// TIA Portal project "Project maybe not work 1.0" (V17) (continued)
REGION Network 7: Step 25 resetting the alarms
   "Data_Block_Reset_Seq".SeqStep[27] := "Data_Block_Reset_Seq".StepNumber = 27;
   "Data_Block_Reset_Seq".SeqConditions[27] := ("Data_Block_Reset_Seq".StepNumber = 27) AND NOT "FS-313.I" AND NOT "FS-214-I" AND "FS-213.I" AND NOT "FS-115.I" AND "FS-114.I" AND NOT "FS-113.I" AND NOT "FS-212.I" AND "HZ-413.I" AND NOT "Fire Alarm" AND NOT "QE-116.I" AND "QE-316.I";
   "Data_Block_Reset_Seq".SeqTimer[27].TON(IN := ("Data_Block_Reset_Seq".StepNumber = 27) AND (("FS-314.I" AND NOT "FS-315.I") OR (NOT "FS-315.I" AND NOT "FS-314.I")) AND NOT "FS-315.I" AND "Data_Block_Reset_Seq".SeqConditions[27],
                           PT := T#50MS);
   IF "Data_Block_Reset_Seq".SeqTimer[27].Q THEN
       "FCS-311.O" := FALSE;
       "FCS-312.O" := TRUE;
   END_IF;
   #_w1 := "Data_Block_Reset_Seq".StepNumber = 27;
   IF "Data_Block_Reset_Seq".SeqTimer[27].Q THEN "Data_Block_Reset_Seq".StepNumber := 28; END_IF;
   "Data_Block_Reset_Seq".SeqTimer_1[89].TON(IN := #_w1 AND NOT "FS-314.I" AND "FS-315.I" AND "Data_Block_Reset_Seq".SeqConditions[27],
                           PT := T#50MS);
   IF "Data_Block_Reset_Seq".SeqTimer_1[89].Q THEN "Data_Block_Reset_Seq".StepNumber := 28; END_IF;
END_REGION

REGION Network 8: Step 25 resetting the alarms
   "Data_Block_Reset_Seq".SeqStep[28] := "Data_Block_Reset_Seq".StepNumber = 28;
   "Data_Block_Reset_Seq".SeqConditions[28] := ("Data_Block_Reset_Seq".StepNumber = 28) AND NOT "FS-314.I" AND "FS-315.I" AND NOT "FS-313.I" AND NOT "FS-214-I" AND "FS-213.I" AND NOT "FS-115.I" AND "FS-114.I" AND NOT "FS-113.I" AND NOT "FS-212.I" AND "HZ-413.I" AND NOT "Fire Alarm" AND NOT "QE-116.I" AND "QE-316.I";
   "Data_Block_Reset_Seq".SeqTimer[28].TON(IN := ("Data_Block_Reset_Seq".StepNumber = 28) AND "Data_Block_Reset_Seq".SeqConditions[28],
                           PT := T#50MS);
   IF "Data_Block_Reset_Seq".SeqTimer[28].Q THEN
       "FCS-312.O" := FALSE;
       "Data_Block_Reset_Seq".StepNumber := 30;
   END_IF;
END_REGION

REGION Network 9: Step 25 resetting the alarms
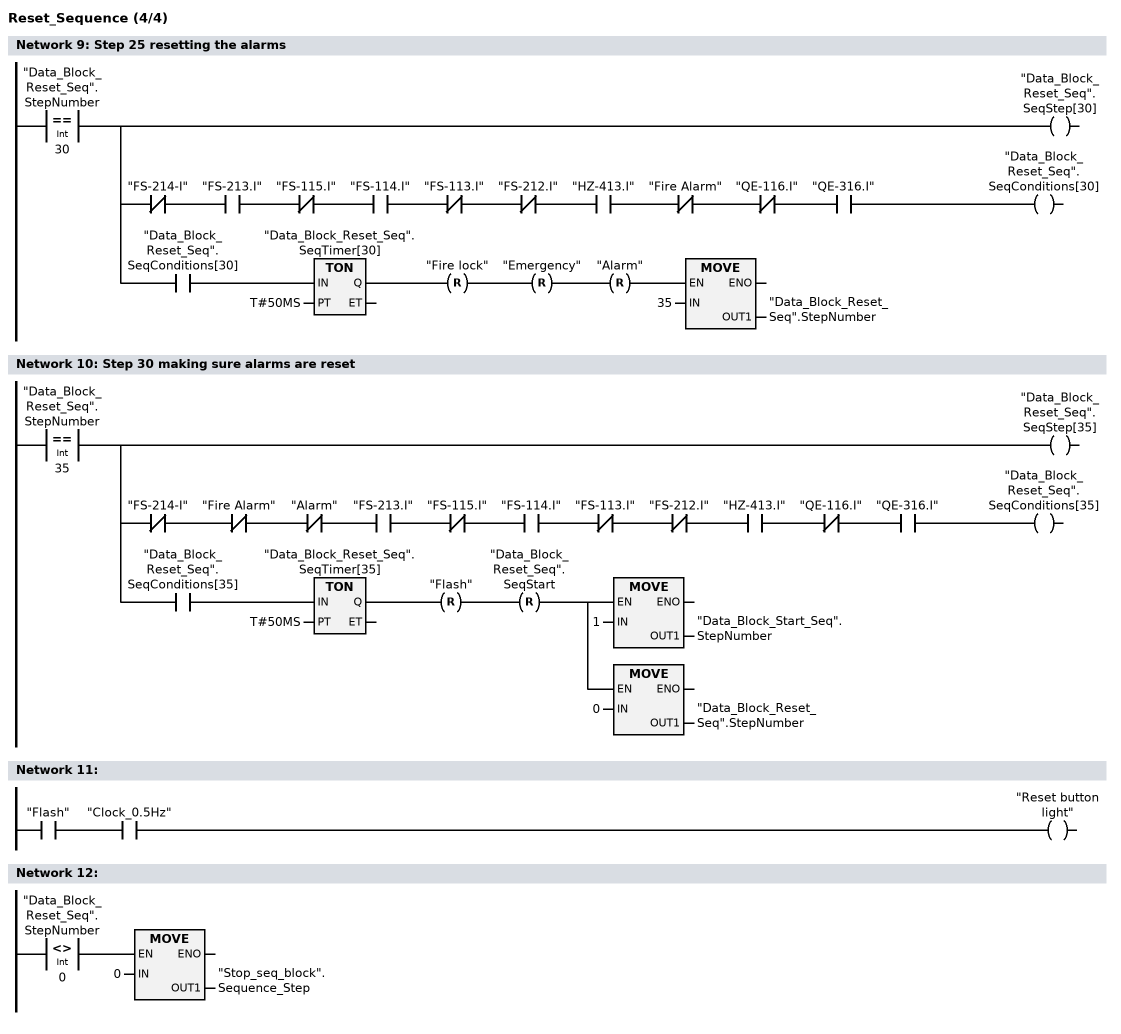
   "Data_Block_Reset_Seq".SeqStep[30] := "Data_Block_Reset_Seq".StepNumber = 30;
   "Data_Block_Reset_Seq".SeqConditions[30] := ("Data_Block_Reset_Seq".StepNumber = 30) AND NOT "FS-214-I" AND "FS-213.I" AND NOT "FS-115.I" AND "FS-114.I" AND NOT "FS-113.I" AND NOT "FS-212.I" AND "HZ-413.I" AND NOT "Fire Alarm" AND NOT "QE-116.I" AND "QE-316.I";
   "Data_Block_Reset_Seq".SeqTimer[30].TON(IN := ("Data_Block_Reset_Seq".StepNumber = 30) AND "Data_Block_Reset_Seq".SeqConditions[30],
                           PT := T#50MS);
   IF "Data_Block_Reset_Seq".SeqTimer[30].Q THEN
       "Fire lock" := FALSE;
       "Emergency" := FALSE;
       "Alarm" := FALSE;
       "Data_Block_Reset_Seq".StepNumber := 35;
   END_IF;
END_REGION

REGION Network 10: Step 30 making sure alarms are reset
   "Data_Block_Reset_Seq".SeqStep[35] := "Data_Block_Reset_Seq".StepNumber = 35;
   "Data_Block_Reset_Seq".SeqConditions[35] := ("Data_Block_Reset_Seq".StepNumber = 35) AND NOT "FS-214-I" AND NOT "Fire Alarm" AND NOT "Alarm" AND "FS-213.I" AND NOT "FS-115.I" AND "FS-114.I" AND NOT "FS-113.I" AND NOT "FS-212.I" AND "HZ-413.I" AND NOT "QE-116.I" AND "QE-316.I";
   "Data_Block_Reset_Seq".SeqTimer[35].TON(IN := ("Data_Block_Reset_Seq".StepNumber = 35) AND "Data_Block_Reset_Seq".SeqConditions[35],
                           PT := T#50MS);
   IF "Data_Block_Reset_Seq".SeqTimer[35].Q THEN
       "Flash" := FALSE;
       "Data_Block_Reset_Seq".SeqStart := FALSE;
       "Data_Block_Start_Seq".StepNumber := 1;
       "Data_Block_Reset_Seq".StepNumber := 0;
   END_IF;
END_REGION

REGION Network 11
   RUNG wire#powerrail
      Contact( "Flash" )
      Contact( "Clock_0.5Hz" )
      Coil( "Reset button light" )
   END_RUNG
   // the same network as SCL:
   "Reset button light" := "Flash" AND "Clock_0.5Hz";
END_REGION

REGION Network 12
   RUNG wire#powerrail
      { S7_Templates := "SrcType := Int" } NE_Contact(in1 := "Data_Block_Reset_Seq".StepNumber, in2 := 0)
      Move(in := 0, out1 => "Stop_seq_block".Sequence_Step)
   END_RUNG
   // the same network as SCL:
   IF "Data_Block_Reset_Seq".StepNumber <> 0 THEN "Stop_seq_block".Sequence_Step := 0; END_IF;
END_REGION
END_FUNCTION

FUNCTION "Stop_Sequence" : Void   // FC2, LAD
{ S7_Optimized_Access := 'TRUE' }
VERSION : 0.1
   VAR_TEMP   // added for the SCL form of the ladder/FBD networks
      _w1 : Bool;
      _w2 : Bool;
   END_VAR
BEGIN

REGION Network 1
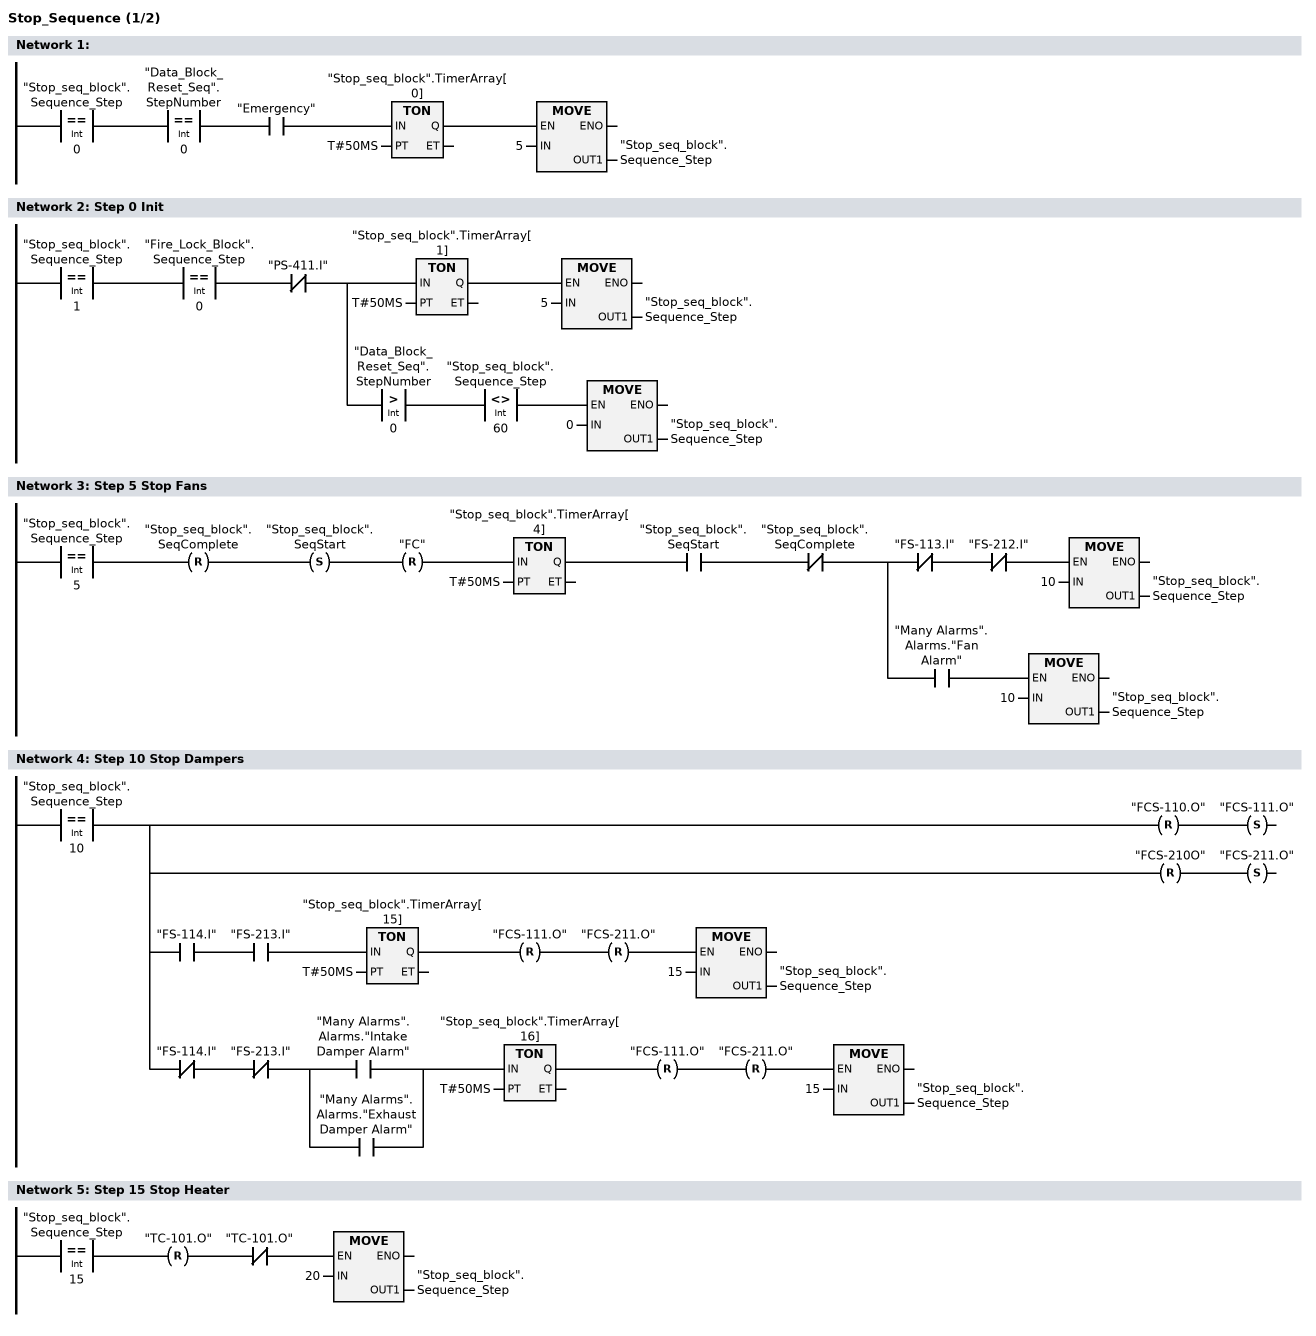
   "Stop_seq_block".TimerArray[0].TON(IN := ("Stop_seq_block".Sequence_Step = 0) AND ("Data_Block_Reset_Seq".StepNumber = 0) AND "Emergency",
                           PT := T#50MS);
   IF "Stop_seq_block".TimerArray[0].Q THEN "Stop_seq_block".Sequence_Step := 5; END_IF;
END_REGION

REGION Network 2: Step 0 Init
   #_w1 := ("Stop_seq_block".Sequence_Step = 1) AND ("Fire_Lock_Block".Sequence_Step = 0) AND NOT "PS-411.I";
   "Stop_seq_block".TimerArray[1].TON(IN := #_w1, PT := T#50MS);
   IF "Stop_seq_block".TimerArray[1].Q THEN "Stop_seq_block".Sequence_Step := 5; END_IF;
   IF #_w1 AND ("Data_Block_Reset_Seq".StepNumber > 0) AND ("Stop_seq_block".Sequence_Step <> 60) THEN
       "Stop_seq_block".Sequence_Step := 0;
   END_IF;
END_REGION

REGION Network 3: Step 5 Stop Fans
   #_w1 := "Stop_seq_block".Sequence_Step = 5;
   IF #_w1 THEN
       "Stop_seq_block".SeqComplete := FALSE;
       "Stop_seq_block".SeqStart := TRUE;
       "FC" := FALSE;
   END_IF;
   "Stop_seq_block".TimerArray[4].TON(IN := #_w1, PT := T#50MS);
   #_w2 := "Stop_seq_block".TimerArray[4].Q AND "Stop_seq_block".SeqStart AND NOT "Stop_seq_block".SeqComplete;
   IF #_w2 AND NOT "FS-113.I" AND NOT "FS-212.I" THEN "Stop_seq_block".Sequence_Step := 10; END_IF;
   IF #_w2 AND "Many Alarms".Alarms."Fan Alarm" THEN "Stop_seq_block".Sequence_Step := 10; END_IF;
END_REGION

REGION Network 4: Step 10 Stop Dampers
   #_w1 := "Stop_seq_block".Sequence_Step = 10;
   IF #_w1 THEN
       "FCS-110.O" := FALSE;
       "FCS-111.O" := TRUE;
       "FCS-210O" := FALSE;
       "FCS-211.O" := TRUE;
   END_IF;
   "Stop_seq_block".TimerArray[15].TON(IN := #_w1 AND "FS-114.I" AND "FS-213.I", PT := T#50MS);
   IF "Stop_seq_block".TimerArray[15].Q THEN
       "FCS-111.O" := FALSE;
       "FCS-211.O" := FALSE;
       "Stop_seq_block".Sequence_Step := 15;
   END_IF;
   "Stop_seq_block".TimerArray[16].TON(IN := #_w1 AND NOT "FS-114.I" AND NOT "FS-213.I" AND ("Many Alarms".Alarms."Intake Damper Alarm" OR "Many Alarms".Alarms."Exhaust Damper Alarm"),
                           PT := T#50MS);
   IF "Stop_seq_block".TimerArray[16].Q THEN
       "FCS-111.O" := FALSE;
       "FCS-211.O" := FALSE;
       "Stop_seq_block".Sequence_Step := 15;
   END_IF;
END_REGION

REGION Network 5: Step 15 Stop Heater
   RUNG wire#powerrail
      { S7_Templates := "SrcType := Int" } EQ_Contact(in1 := "Stop_seq_block".Sequence_Step, in2 := 15)
      R_Coil( "TC-101.O" )
      I_Contact( "TC-101.O" )
      Move(in := 20, out1 => "Stop_seq_block".Sequence_Step)
   END_RUNG
   // the same network as SCL:
   #_w1 := "Stop_seq_block".Sequence_Step = 15;
   IF #_w1 THEN "TC-101.O" := FALSE; END_IF;
   IF #_w1 AND NOT "TC-101.O" THEN "Stop_seq_block".Sequence_Step := 20; END_IF;
END_REGION

REGION Network 6: Step 20 Sequence Complete
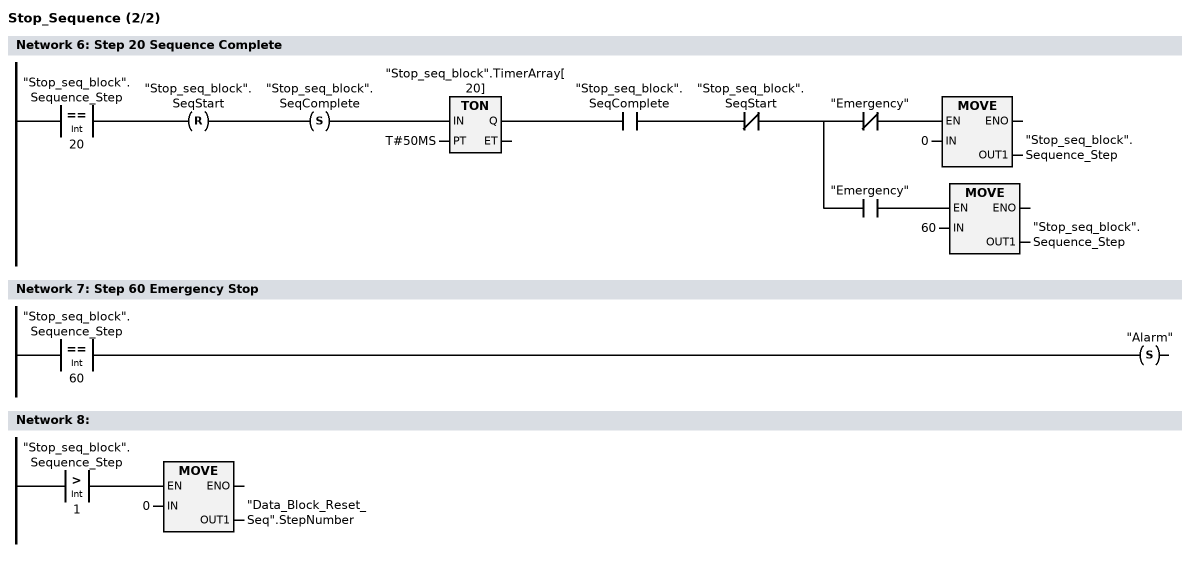
   #_w1 := "Stop_seq_block".Sequence_Step = 20;
   IF #_w1 THEN
       "Stop_seq_block".SeqStart := FALSE;
       "Stop_seq_block".SeqComplete := TRUE;
   END_IF;
   "Stop_seq_block".TimerArray[20].TON(IN := #_w1, PT := T#50MS);
   #_w2 := "Stop_seq_block".TimerArray[20].Q AND "Stop_seq_block".SeqComplete AND NOT "Stop_seq_block".SeqStart;
   IF #_w2 AND NOT "Emergency" THEN "Stop_seq_block".Sequence_Step := 0; END_IF;
   IF #_w2 AND "Emergency" THEN "Stop_seq_block".Sequence_Step := 60; END_IF;
END_REGION

REGION Network 7: Step 60 Emergency Stop
   RUNG wire#powerrail
      { S7_Templates := "SrcType := Int" } EQ_Contact(in1 := "Stop_seq_block".Sequence_Step, in2 := 60)
      S_Coil( "Alarm" )
   END_RUNG
   // the same network as SCL:
   IF "Stop_seq_block".Sequence_Step = 60 THEN "Alarm" := TRUE; END_IF;
END_REGION

REGION Network 8
   RUNG wire#powerrail
      { S7_Templates := "SrcType := Int" } GT_Contact(in1 := "Stop_seq_block".Sequence_Step, in2 := 1)
      Move(in := 0, out1 => "Data_Block_Reset_Seq".StepNumber)
   END_RUNG
   // the same network as SCL:
   IF "Stop_seq_block".Sequence_Step > 1 THEN "Data_Block_Reset_Seq".StepNumber := 0; END_IF;
END_REGION
END_FUNCTION

FUNCTION "Fire_Lock_Sequence" : Void   // FC3, LAD
{ S7_Optimized_Access := 'TRUE' }
VERSION : 0.1
   VAR_TEMP   // added for the SCL form of the ladder/FBD networks
      _w1 : Bool;
      _w2 : Bool;
   END_VAR
BEGIN

REGION Network 1
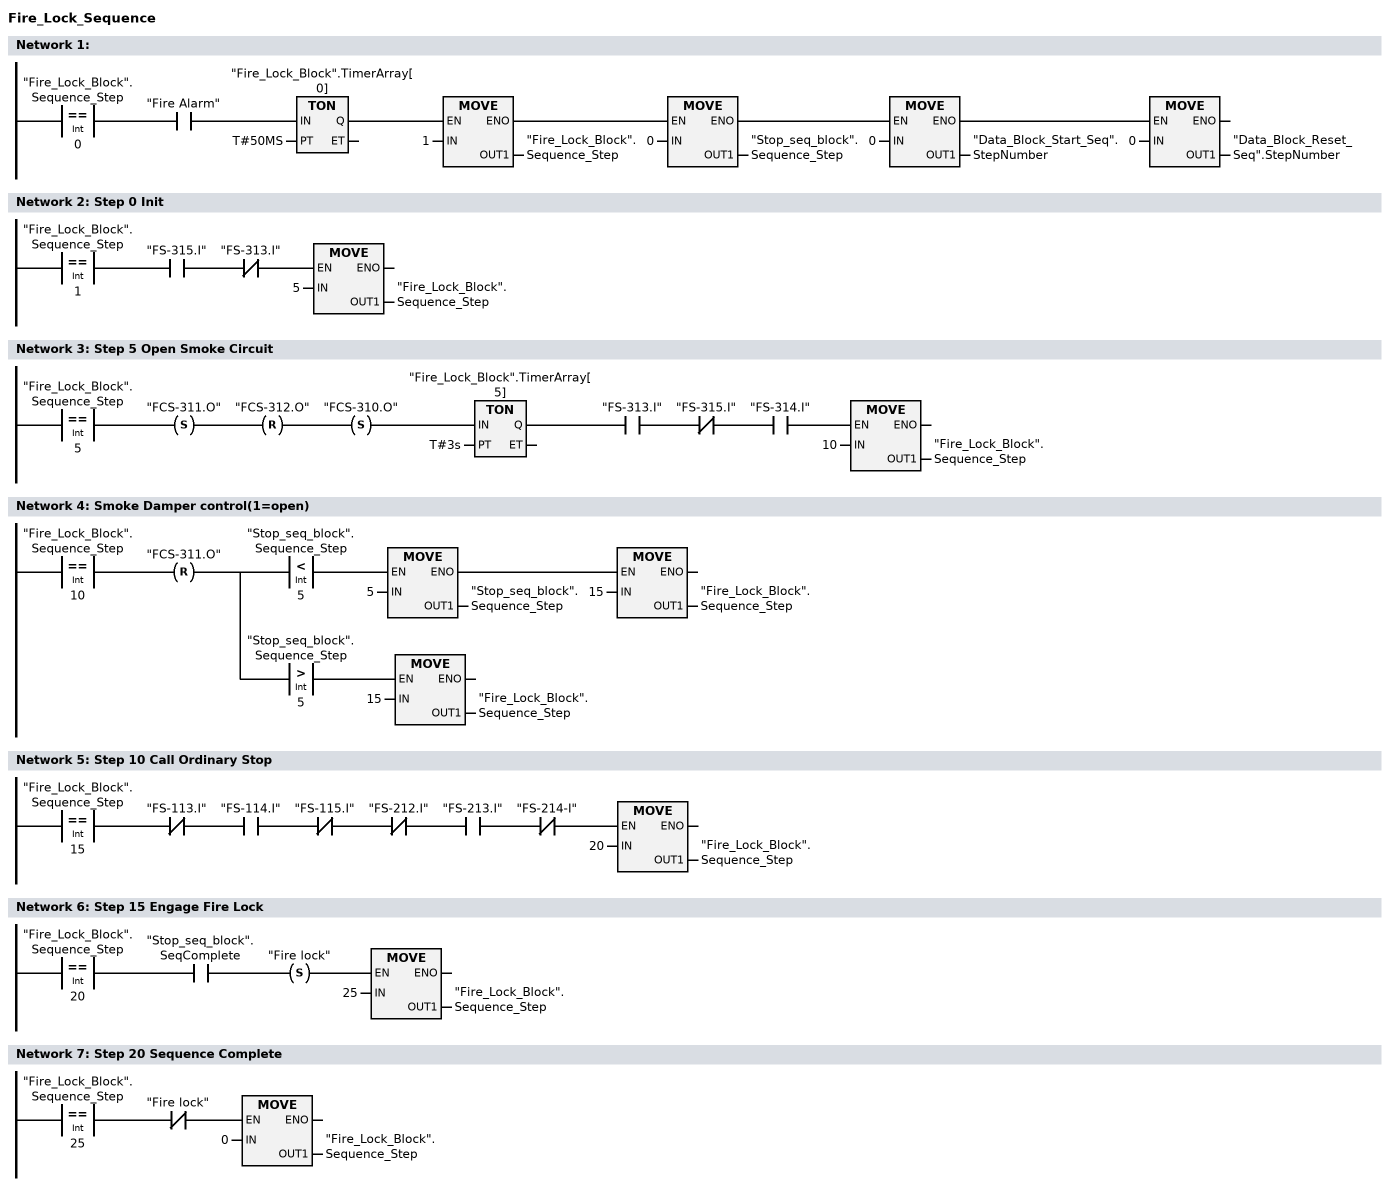
   "Fire_Lock_Block".TimerArray[0].TON(IN := ("Fire_Lock_Block".Sequence_Step = 0) AND "Fire Alarm",
                           PT := T#50MS);
   IF "Fire_Lock_Block".TimerArray[0].Q THEN
       "Fire_Lock_Block".Sequence_Step := 1;
       "Stop_seq_block".Sequence_Step := 0;
       "Data_Block_Start_Seq".StepNumber := 0;
       "Data_Block_Reset_Seq".StepNumber := 0;
   END_IF;
END_REGION

REGION Network 2: Step 0 Init
   RUNG wire#powerrail
      { S7_Templates := "SrcType := Int" } EQ_Contact(in1 := "Fire_Lock_Block".Sequence_Step, in2 := 1)
      Contact( "FS-315.I" )
      I_Contact( "FS-313.I" )
      Move(in := 5, out1 => "Fire_Lock_Block".Sequence_Step)
   END_RUNG
   // the same network as SCL:
   IF ("Fire_Lock_Block".Sequence_Step = 1) AND "FS-315.I" AND NOT "FS-313.I" THEN
       "Fire_Lock_Block".Sequence_Step := 5;
   END_IF;
END_REGION

REGION Network 3: Step 5 Open Smoke Circuit
   #_w1 := "Fire_Lock_Block".Sequence_Step = 5;
   IF #_w1 THEN
       "FCS-311.O" := TRUE;
       "FCS-312.O" := FALSE;
       "FCS-310.O" := TRUE;
   END_IF;
   "Fire_Lock_Block".TimerArray[5].TON(IN := #_w1, PT := T#3s);
   IF "Fire_Lock_Block".TimerArray[5].Q AND "FS-313.I" AND NOT "FS-315.I" AND "FS-314.I" THEN
       "Fire_Lock_Block".Sequence_Step := 10;
   END_IF;
END_REGION

REGION Network 4: Smoke Damper control(1=open)
   RUNG wire#powerrail
      { S7_Templates := "SrcType := Int" } EQ_Contact(in1 := "Fire_Lock_Block".Sequence_Step, in2 := 10)
      R_Coil( "FCS-311.O" )
      wire#w1
      { S7_Templates := "SrcType := Int" } LT_Contact(in1 := "Stop_seq_block".Sequence_Step, in2 := 5)
      Move(in := 5, out1 => "Stop_seq_block".Sequence_Step)
      Move(in := 15, out1 => "Fire_Lock_Block".Sequence_Step)
   END_RUNG
   RUNG wire#w1
      { S7_Templates := "SrcType := Int" } GT_Contact(in1 := "Stop_seq_block".Sequence_Step, in2 := 5)
      Move(in := 15, out1 => "Fire_Lock_Block".Sequence_Step)
   END_RUNG
   // the same network as SCL:
   #_w1 := "Fire_Lock_Block".Sequence_Step = 10;
   IF #_w1 THEN "FCS-311.O" := FALSE; END_IF;
   #_w2 := #_w1 AND ("Stop_seq_block".Sequence_Step < 5);
   IF #_w2 THEN
       "Stop_seq_block".Sequence_Step := 5;
       "Fire_Lock_Block".Sequence_Step := 15;
   END_IF;
   IF #_w1 AND ("Stop_seq_block".Sequence_Step > 5) THEN "Fire_Lock_Block".Sequence_Step := 15; END_IF;
END_REGION

REGION Network 5: Step 10 Call Ordinary Stop
   RUNG wire#powerrail
      { S7_Templates := "SrcType := Int" } EQ_Contact(in1 := "Fire_Lock_Block".Sequence_Step, in2 := 15)
      I_Contact( "FS-113.I" )
      Contact( "FS-114.I" )
      I_Contact( "FS-115.I" )
      I_Contact( "FS-212.I" )
      Contact( "FS-213.I" )
      I_Contact( "FS-214-I" )
      Move(in := 20, out1 => "Fire_Lock_Block".Sequence_Step)
   END_RUNG
   // the same network as SCL:
   IF ("Fire_Lock_Block".Sequence_Step = 15) AND NOT "FS-113.I" AND "FS-114.I" AND NOT "FS-115.I" AND NOT "FS-212.I" AND "FS-213.I" AND NOT "FS-214-I" THEN
       "Fire_Lock_Block".Sequence_Step := 20;
   END_IF;
END_REGION

REGION Network 6: Step 15 Engage Fire Lock
   RUNG wire#powerrail
      { S7_Templates := "SrcType := Int" } EQ_Contact(in1 := "Fire_Lock_Block".Sequence_Step, in2 := 20)
      Contact( "Stop_seq_block".SeqComplete )
      S_Coil( "Fire lock" )
      Move(in := 25, out1 => "Fire_Lock_Block".Sequence_Step)
   END_RUNG
   // the same network as SCL:
   IF ("Fire_Lock_Block".Sequence_Step = 20) AND "Stop_seq_block".SeqComplete THEN
       "Fire lock" := TRUE;
       "Fire_Lock_Block".Sequence_Step := 25;
   END_IF;
END_REGION

REGION Network 7: Step 20 Sequence Complete
   RUNG wire#powerrail
      { S7_Templates := "SrcType := Int" } EQ_Contact(in1 := "Fire_Lock_Block".Sequence_Step, in2 := 25)
      I_Contact( "Fire lock" )
      Move(in := 0, out1 => "Fire_Lock_Block".Sequence_Step)
   END_RUNG
   // the same network as SCL:
   IF ("Fire_Lock_Block".Sequence_Step = 25) AND NOT "Fire lock" THEN
       "Fire_Lock_Block".Sequence_Step := 0;
   END_IF;
END_REGION

REGION Network 8: Step 60 Hardware Error
END_REGION
END_FUNCTION

FUNCTION "Start_Sequence" : Void   // FC11, LAD
{ S7_Optimized_Access := 'TRUE' }
VERSION : 0.1
   VAR_TEMP   // added for the SCL form of the ladder/FBD networks
      _w1 : Bool;
      _w2 : Bool;
   END_VAR
BEGIN

REGION Network 1
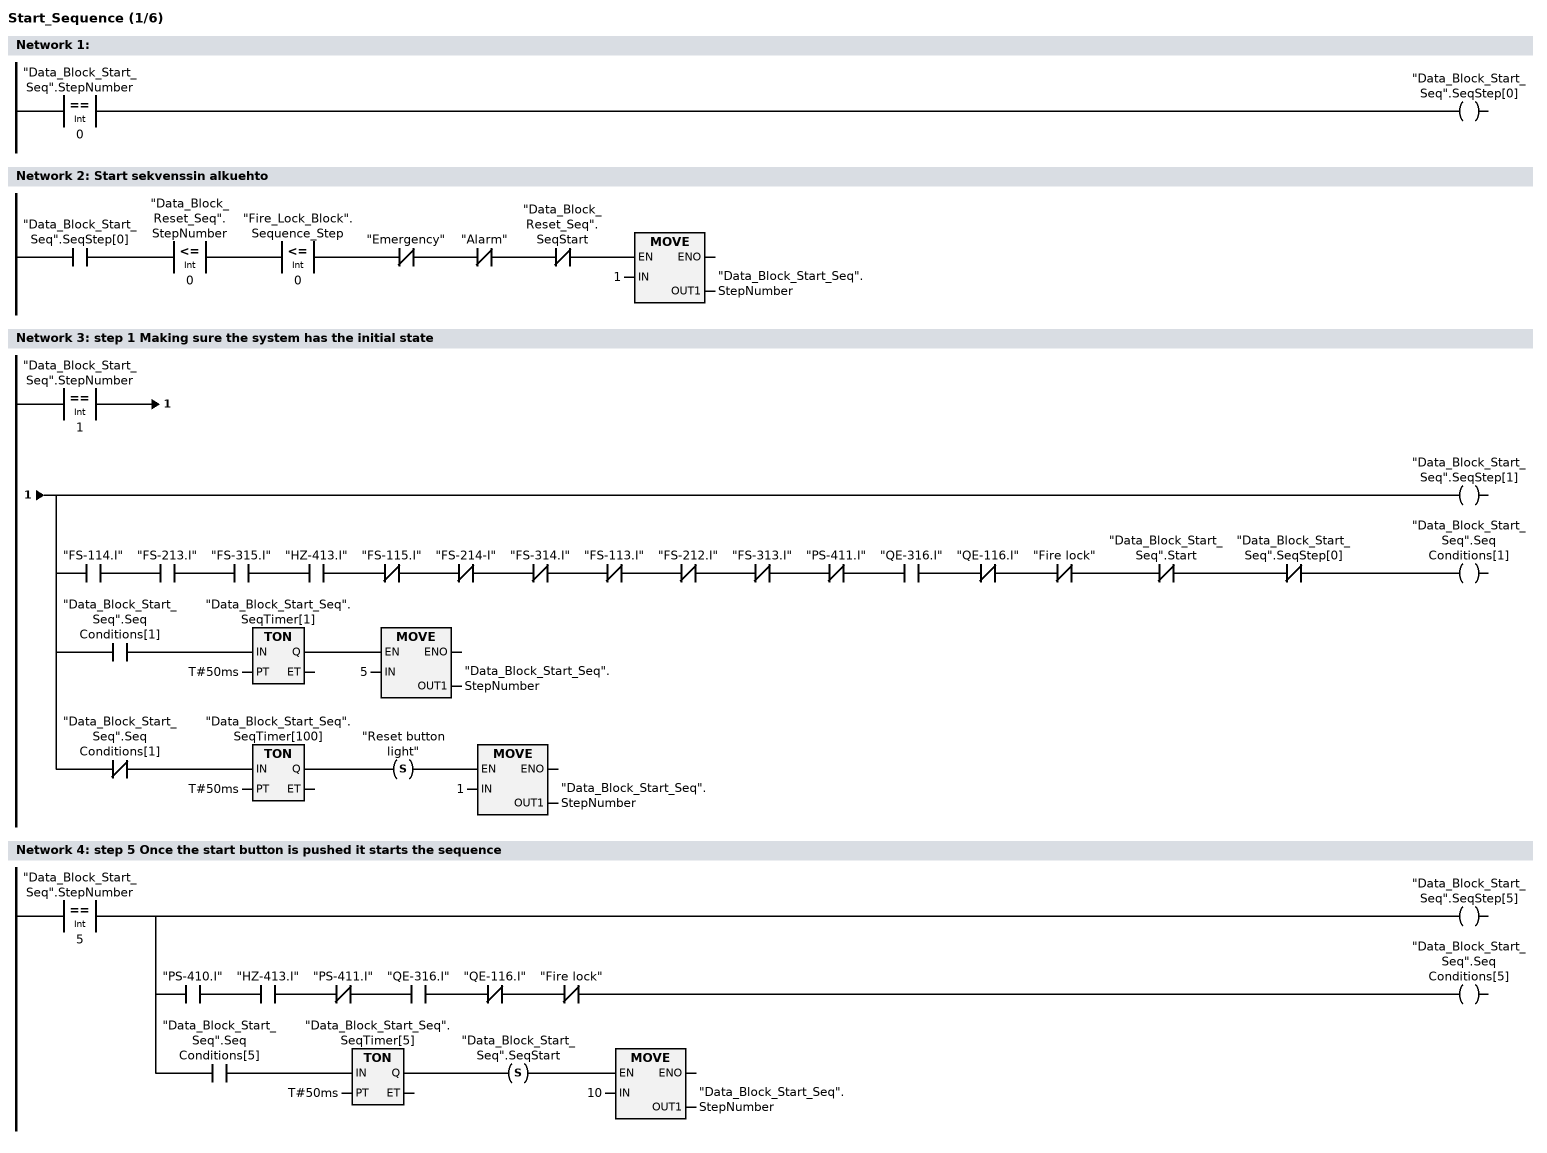
   RUNG wire#powerrail
      { S7_Templates := "SrcType := Int" } EQ_Contact(in1 := "Data_Block_Start_Seq".StepNumber, in2 := 0)
      Coil( "Data_Block_Start_Seq".SeqStep[0] )
   END_RUNG
   // the same network as SCL:
   "Data_Block_Start_Seq".SeqStep[0] := "Data_Block_Start_Seq".StepNumber = 0;
END_REGION

REGION Network 2: Start sekvenssin alkuehto
   RUNG wire#powerrail
      Contact( "Data_Block_Start_Seq".SeqStep[0] )
      { S7_Templates := "SrcType := Int" } LE_Contact(in1 := "Data_Block_Reset_Seq".StepNumber, in2 := 0)
      { S7_Templates := "SrcType := Int" } LE_Contact(in1 := "Fire_Lock_Block".Sequence_Step, in2 := 0)
      I_Contact( "Emergency" )
      I_Contact( "Alarm" )
      I_Contact( "Data_Block_Reset_Seq".SeqStart )
      Move(in := 1, out1 => "Data_Block_Start_Seq".StepNumber)
   END_RUNG
   // the same network as SCL:
   IF "Data_Block_Start_Seq".SeqStep[0] AND ("Data_Block_Reset_Seq".StepNumber <= 0) AND ("Fire_Lock_Block".Sequence_Step <= 0) AND NOT "Emergency" AND NOT "Alarm" AND NOT "Data_Block_Reset_Seq".SeqStart THEN
       "Data_Block_Start_Seq".StepNumber := 1;
   END_IF;
END_REGION

REGION Network 3: step 1 Making sure the system has the initial state
   "Data_Block_Start_Seq".SeqStep[1] := "Data_Block_Start_Seq".StepNumber = 1;
   "Data_Block_Start_Seq".SeqConditions[1] := ("Data_Block_Start_Seq".StepNumber = 1) AND "FS-114.I" AND "FS-213.I" AND "FS-315.I" AND "HZ-413.I" AND NOT "FS-115.I" AND NOT "FS-214-I" AND NOT "FS-314.I" AND NOT "FS-113.I" AND NOT "FS-212.I" AND NOT "FS-313.I" AND NOT "PS-411.I" AND "QE-316.I" AND NOT "QE-116.I" AND NOT "Fire lock" AND NOT "Data_Block_Start_Seq".Start AND NOT "Data_Block_Start_Seq".SeqStep[0];
   "Data_Block_Start_Seq".SeqTimer[1].TON(IN := ("Data_Block_Start_Seq".StepNumber = 1) AND "Data_Block_Start_Seq".SeqConditions[1],
                           PT := T#50ms);
   #_w1 := "Data_Block_Start_Seq".StepNumber = 1;
   IF "Data_Block_Start_Seq".SeqTimer[1].Q THEN "Data_Block_Start_Seq".StepNumber := 5; END_IF;
   "Data_Block_Start_Seq".SeqTimer[100].TON(IN := #_w1 AND NOT "Data_Block_Start_Seq".SeqConditions[1],
                           PT := T#50ms);
   IF "Data_Block_Start_Seq".SeqTimer[100].Q THEN
       "Reset button light" := TRUE;
       "Data_Block_Start_Seq".StepNumber := 1;
   END_IF;
END_REGION

REGION Network 4: step 5 Once the start button is pushed it starts the sequence
   "Data_Block_Start_Seq".SeqStep[5] := "Data_Block_Start_Seq".StepNumber = 5;
   "Data_Block_Start_Seq".SeqConditions[5] := ("Data_Block_Start_Seq".StepNumber = 5) AND "PS-410.I" AND "HZ-413.I" AND NOT "PS-411.I" AND "QE-316.I" AND NOT "QE-116.I" AND NOT "Fire lock";
   "Data_Block_Start_Seq".SeqTimer[5].TON(IN := ("Data_Block_Start_Seq".StepNumber = 5) AND "Data_Block_Start_Seq".SeqConditions[5],
                           PT := T#50ms);
   IF "Data_Block_Start_Seq".SeqTimer[5].Q THEN
       "Data_Block_Start_Seq".SeqStart := TRUE;
       "Data_Block_Start_Seq".StepNumber := 10;
   END_IF;
END_REGION

REGION Network 5: step 10 Makes sure the start sequence has been started after which it starts to open the dampers. Also makes sure the closing control is released.
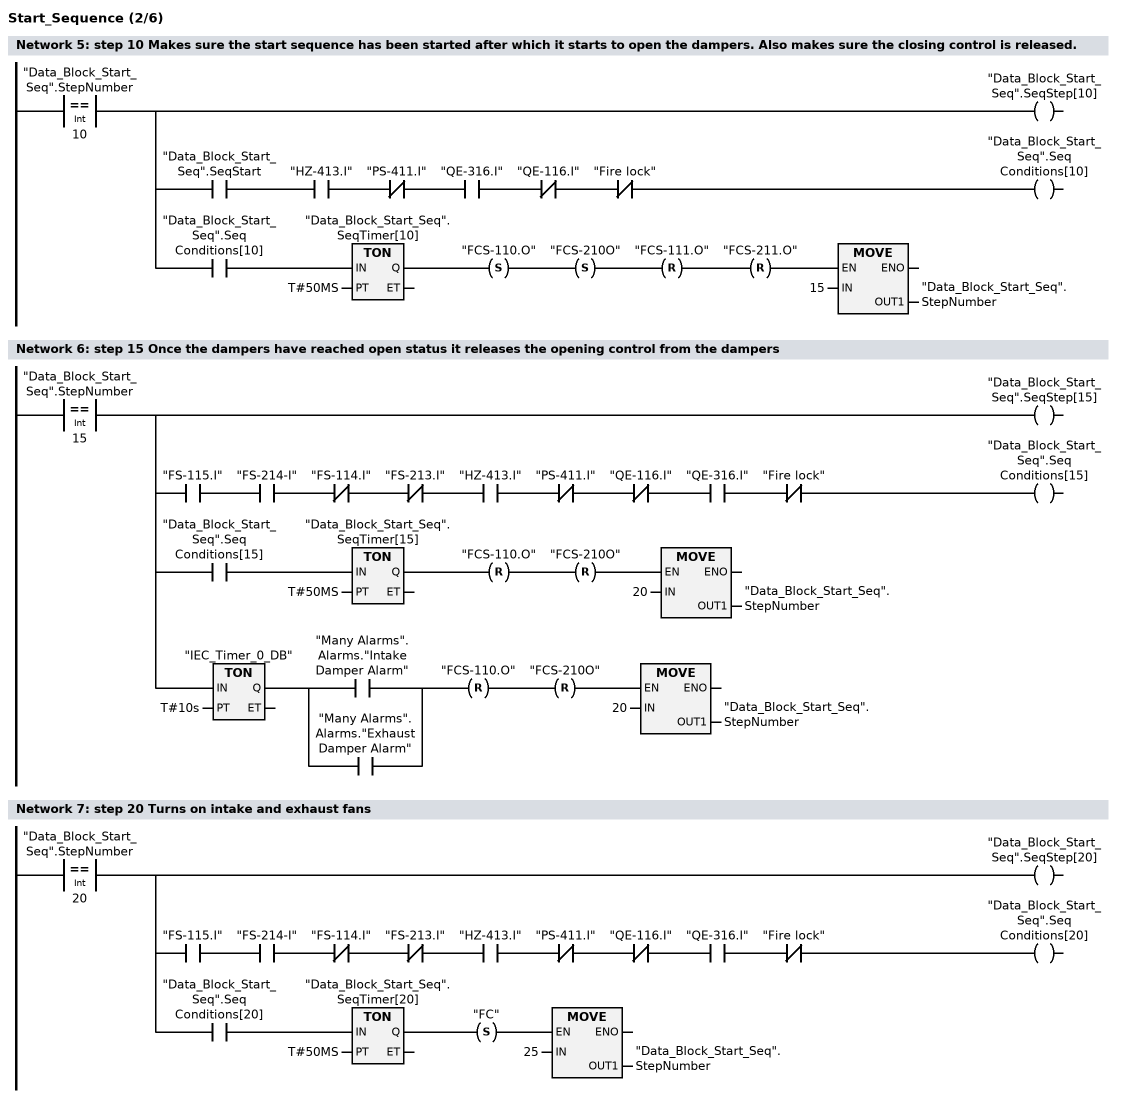
   "Data_Block_Start_Seq".SeqStep[10] := "Data_Block_Start_Seq".StepNumber = 10;
   "Data_Block_Start_Seq".SeqConditions[10] := ("Data_Block_Start_Seq".StepNumber = 10) AND "Data_Block_Start_Seq".SeqStart AND "HZ-413.I" AND NOT "PS-411.I" AND "QE-316.I" AND NOT "QE-116.I" AND NOT "Fire lock";
   "Data_Block_Start_Seq".SeqTimer[10].TON(IN := ("Data_Block_Start_Seq".StepNumber = 10) AND "Data_Block_Start_Seq".SeqConditions[10],
                           PT := T#50MS);
   IF "Data_Block_Start_Seq".SeqTimer[10].Q THEN
       "FCS-110.O" := TRUE;
       "FCS-210O" := TRUE;
       "FCS-111.O" := FALSE;
       "FCS-211.O" := FALSE;
       "Data_Block_Start_Seq".StepNumber := 15;
   END_IF;
END_REGION

REGION Network 6: step 15 Once the dampers have reached open status it releases the opening control from the dampers
   "Data_Block_Start_Seq".SeqStep[15] := "Data_Block_Start_Seq".StepNumber = 15;
   "Data_Block_Start_Seq".SeqConditions[15] := ("Data_Block_Start_Seq".StepNumber = 15) AND "FS-115.I" AND "FS-214-I" AND NOT "FS-114.I" AND NOT "FS-213.I" AND "HZ-413.I" AND NOT "PS-411.I" AND NOT "QE-116.I" AND "QE-316.I" AND NOT "Fire lock";
   "Data_Block_Start_Seq".SeqTimer[15].TON(IN := ("Data_Block_Start_Seq".StepNumber = 15) AND "Data_Block_Start_Seq".SeqConditions[15],
                           PT := T#50MS);
   IF "Data_Block_Start_Seq".SeqTimer[15].Q THEN
       "FCS-110.O" := FALSE;
       "FCS-210O" := FALSE;
   END_IF;
   #_w1 := "Data_Block_Start_Seq".StepNumber = 15;
   IF "Data_Block_Start_Seq".SeqTimer[15].Q THEN "Data_Block_Start_Seq".StepNumber := 20; END_IF;
   "IEC_Timer_0_DB".TON(IN := #_w1, PT := T#10s);
   IF "IEC_Timer_0_DB".Q AND ("Many Alarms".Alarms."Intake Damper Alarm" OR "Many Alarms".Alarms."Exhaust Damper Alarm") THEN
       "FCS-110.O" := FALSE;
       "FCS-210O" := FALSE;
       "Data_Block_Start_Seq".StepNumber := 20;
   END_IF;
END_REGION
